   "Carrier_51_G120DStatusWord.0" AT %I2912.0 : Bool;   // Bit_00_READY_RUN
   "Carrier_51_G120DStatusWord.1" AT %I2912.1 : Bool;   // Bit_01_READY_ON
   "Carrier_51_G120DStatusWord.2" AT %I2912.2 : Bool;   // Bit_02_ENABLE
   "Carrier_51_G120DStatusWord.3" AT %I2912.3 : Bool;   // Bit_03_FAULT
   "Carrier_51_G120DStatusWord.4" AT %I2912.4 : Bool;   // Bit_04_OFF2
   "Carrier_51_G120DStatusWord.5" AT %I2912.5 : Bool;   // Bit_05_OFF3
   "Carrier_51_G120DStatusWord.6" AT %I2912.6 : Bool;   // Bit_06_LOCK_OUT
   "Carrier_51_G120DStatusWord.7" AT %I2912.7 : Bool;   // Bit_07_WARN
   "Carrier_51_G120DStatusWord.8" AT %I2913.0 : Bool;   // Bit_08_NO_DEVIATION
   "Carrier_51_G120DStatusWord.9" AT %I2913.1 : Bool;   // Bit_09_CONTR_PLC
   "Carrier_51_G120DStatusWord.10" AT %I2913.2 : Bool;   // Bit_10_F_MAX
   "Carrier_51_G120DStatusWord.11" AT %I2913.3 : Bool;   // Bit_11_LIMIT_REACHED
   "Carrier_51_G120DStatusWord.12" AT %I2913.4 : Bool;   // Bit_12_BRAKE_OPEN
   "Carrier_51_G120DStatusWord.13" AT %I2913.5 : Bool;   // Bit_13_NO_OVERTEMP
   "Carrier_51_G120DStatusWord.14" AT %I2913.6 : Bool;   // Bit_14_CW_CCW
   "Carrier_51_G120DStatusWord.15" AT %I2913.7 : Bool;   // Bit_15_OVERL
   "Carrier_51_Slot2_Input" AT %IW2914 : Word;   // SLOT 2 INPUT WORD
   "Carrier_51_CrashDetectSW" AT %I2914.0 : Bool;   // CRASH DETECT SW
   "Carrier_51_SpareSafetyInput(2_1)" AT %I2914.1 : Bool;   // SPARE SAFETY INPUT
   "Carrier_51_SpareSafetyInput(2_2)" AT %I2914.2 : Bool;   // SPARE SAFETY INPUT
   "Carrier_51_SpareSafetyInput(2_3)" AT %I2914.3 : Bool;   // SPARE SAFETY INPUT
   "Carrier_51_SpareSafetyInput(2_4)" AT %I2914.4 : Bool;   // SPARE SAFETY INPUT
   "Carrier_51_SpareSafetyInput(2_5)" AT %I2914.5 : Bool;   // SPARE SAFETY INPUT
   "Carrier_51_SpareSafetyInput(2_6)" AT %I2914.6 : Bool;   // SPARE SAFETY INPUT
   "Carrier_51_SpareSafetyInput(2_7)" AT %I2914.7 : Bool;   // SPARE SAFETY INPUT
   "Carrier_51_Slot3_SafetyOutput" AT %IW2915 : Word;   // SLOT 3 SAFETY OUTPUT WORD
   "Carrier_51_Crash_Detect_OK" AT %I2915.0 : Bool;   // CARRIER CRASH DETECT
   "Carrier_51_SpareSafetyOutput(3_1)" AT %I2915.1 : Bool;   // SPARE SAFETY OUTPUT
   "Carrier_51_SpareSafetyOutput(3_2)" AT %I2915.2 : Bool;   // SPARE SAFETY OUTPUT
   "Carrier_51_SpareSafetyOutput(3_3)" AT %I2915.3 : Bool;   // SPARE SAFETY OUTPUT
   "Carrier_51_SpareSafetyOutput(3_4)" AT %I2915.4 : Bool;   // SPARE SAFETY OUTPUT
   "Carrier_51_SpareSafetyOutput(3_5)" AT %I2915.5 : Bool;   // SPARE SAFETY OUTPUT
   "Carrier_51_SpareSafetyOutput(3_6)" AT %I2915.6 : Bool;   // SPARE SAFETY OUTPUT
   "Carrier_51_SpareSafetyOutput(3_7)" AT %I2915.7 : Bool;   // SPARE SAFETY OUTPUT
   "Carrier_51_Slot4_Input" AT %IW2916 : Word;   // SLOT 4 INPUT WORD
   "Carrier_51_480VPowerOn_MDCB1" AT %I2916.0 : Bool;   // 480 VAC POWER ON MDCB 1
   "Carrier_51_SpareInput(4_1)" AT %I2916.1 : Bool;   // SPARE INPUT
   "Carrier_51_SpareInput(4_2)" AT %I2916.2 : Bool;   // SPARE INPUT
   "Carrier_51_SitopSelectStatus" AT %I2916.3 : Bool;   // SITOP SELECT STATUS
   "Carrier_51_DCsupplyOnPSCB2" AT %I2916.4 : Bool;   // DC SUPPLY ON PSCB 2
   "Carrier_51_SpareInput(4_5)" AT %I2916.5 : Bool;   // SPARE INPUT
   "Carrier_51_SpareInput(4_6)" AT %I2916.6 : Bool;   // SPARE INPUT
   "Carrier_51_SpareInput(4_7)" AT %I2916.7 : Bool;   // SPARE INPUT
   "Carrier_51_PB1_ProdHoldLH" AT %I2917.0 : Bool;   // PB 1 PRODUCTION HOLD LH
   "Carrier_51_PB2_ResetLH" AT %I2917.1 : Bool;   // PB 2 RESET LH
   "Carrier_51_PB3_ProdHoldRH" AT %I2917.2 : Bool;   // PB 3 PRODUCTION HOLD RH
   "Carrier_51_PB4_ResetRH" AT %I2917.3 : Bool;   // PB 4 RESET RH
   "Carrier_51_SpareInput(4_14)" AT %I2917.4 : Bool;   // SPARE INPUT
   "Carrier_51_SpareInput(4_15)" AT %I2917.5 : Bool;   // SPARE INPUT
   "Carrier_51_SpareInput(4_16)" AT %I2917.6 : Bool;   // SPARE INPUT
   "Carrier_51_SpareInput(4_17)" AT %I2917.7 : Bool;   // SPARE INPUT
   "Carrier_51_Slot5_Output" AT %IW2918 : Word;   // SLOT 5 OUTPUT WORD
   "Carrier_51_IRD400_HMI_24VDC_ENABLE" AT %I2918.0 : Bool;   // IRD 400 PANEL HMI 24V DC POWER
   "Carrier_51_FaultLight_LH" AT %I2918.1 : Bool;   // FAULT LIGHT LH
   "Carrier_51_RunLight_LH" AT %I2918.2 : Bool;   // RUN LIGHT LH
   "Carrier_51_FaultLight_RH" AT %I2918.3 : Bool;   // FAULT LIGHT RH
   "Carrier_51_RunLight_RH" AT %I2918.4 : Bool;   // RUN LIGHT RH
   "Carrier_51_SpareOutput(5_5)" AT %I2918.5 : Bool;   // SPARE OUTPUT
   "Carrier_51_SpareOutput(5_6)" AT %I2918.6 : Bool;   // SPARE OUTPUT
   "Carrier_51_SpareOutput(5_7)" AT %I2918.7 : Bool;   // SPARE OUTPUT
   "Carrier_51_ActualSpeed" AT %IW2920 : Word;   // ACTUAL SPEED
   "Carrier_51_CarrierDriveAlarm" AT %IW2922 : Word;   // CARRIER DRIVE ALARM
   "Carrier_51_CarrierDriveWarning" AT %IW2924 : Word;   // CARRIER DRIVE WARNING
   "Carrier_52_Status" AT %IW2950 : Word;   // CARRIER STATUS WORD
   "Carrier_52_Status.0" AT %I2950.0 : Bool;   // HEARTBEAT
   "Carrier_52_Status.1" AT %I2950.1 : Bool;   // MANUAL
   "Carrier_52_Status.2" AT %I2950.2 : Bool;   // IN_AUTO
   "Carrier_52_Status.3" AT %I2950.3 : Bool;   // POSITIONING_COMPLETE
   "Carrier_52_Status.4" AT %I2950.4 : Bool;   // PRODUCTION HOLD
   "Carrier_52_Status.5" AT %I2950.5 : Bool;   // CARRIER MOVING FORWARD
   "Carrier_52_Status.6" AT %I2950.6 : Bool;   // CARRIER MOVING REVERSE
   "Carrier_52_Status.7" AT %I2950.7 : Bool;   // CARRIER FAULT
   "Carrier_52_Status.8" AT %I2951.0 : Bool;   // CRASH DETECT TRIPPED
   "Carrier_52_Status.9" AT %I2951.1 : Bool;
   "Carrier_52_Status.10" AT %I2951.2 : Bool;
   "Carrier_52_Status.11" AT %I2951.3 : Bool;
   "Carrier_52_Status.12" AT %I2951.4 : Bool;
   "Carrier_52_Status.13" AT %I2951.5 : Bool;
   "Carrier_52_Status.14" AT %I2951.6 : Bool;
   "Carrier_52_Status.15" AT %I2951.7 : Bool;
   "Carrier_52_SDCFaultCode" AT %IW2952 : Word;   // SDC FAULT CODE
   "Carrier_52_CarrierPosition" AT %ID2954 : DWord;   // CARRIER POSITION
   "Carrier_52_CarrierNumber" AT %IW2958 : Word;   // CARRIER NUMBER
   "Carrier_52_G120DControlWord" AT %IW2960 : Word;   // G120D_STW1_CONTROL
   "Carrier_52_G120DControlWord.0" AT %I2960.0 : Bool;   // Bit_00_ON
   "Carrier_52_G120DControlWord.1" AT %I2960.1 : Bool;   // Bit_01_AUS2_INH
   "Carrier_52_G120DControlWord.2" AT %I2960.2 : Bool;   // Bit_02_AUS3_STOP
   "Carrier_52_G120DControlWord.3" AT %I2960.3 : Bool;   // Bit_03_EN
   "Carrier_52_G120DControlWord.4" AT %I2960.4 : Bool;   // Bit_04_EN_RAMP
   "Carrier_52_G120DControlWord.5" AT %I2960.5 : Bool;   // Bit_05_START_RAMP
   "Carrier_52_G120DControlWord.6" AT %I2960.6 : Bool;   // Bit_06_SETPOINT
   "Carrier_52_G120DControlWord.7" AT %I2960.7 : Bool;   // Bit_07_RESET
   "Carrier_52_G120DControlWord.8" AT %I2961.0 : Bool;   // Bit_08_JOG_R
   "Carrier_52_G120DControlWord.9" AT %I2961.1 : Bool;   // Bit_09_JOG_L
   "Carrier_52_G120DControlWord.10" AT %I2961.2 : Bool;   // Bit_10_CONTR_PLC
   "Carrier_52_G120DControlWord.11" AT %I2961.3 : Bool;   // Bit_11_REVERSE
   "Carrier_52_G120DControlWord.12" AT %I2961.4 : Bool;   // Bit_12_BRAKE_RELEASE
   "Carrier_52_G120DControlWord.13" AT %I2961.5 : Bool;   // Bit_13_DDS
   "Carrier_52_G120DControlWord.14" AT %I2961.6 : Bool;   // Bit_14_DO0
   "Carrier_52_G120DControlWord.15" AT %I2961.7 : Bool;   // Bit_15_DO1
   "Carrier_52_G120DStatusWord" AT %IW2962 : Word;   // G120D_ZSW1_STATUS
   "Carrier_52_G120DStatusWord.0" AT %I2962.0 : Bool;   // Bit_00_READY_RUN
   "Carrier_52_G120DStatusWord.1" AT %I2962.1 : Bool;   // Bit_01_READY_ON
   "Carrier_52_G120DStatusWord.2" AT %I2962.2 : Bool;   // Bit_02_ENABLE
   "Carrier_52_G120DStatusWord.3" AT %I2962.3 : Bool;   // Bit_03_FAULT
   "Carrier_52_G120DStatusWord.4" AT %I2962.4 : Bool;   // Bit_04_OFF2
   "Carrier_52_G120DStatusWord.5" AT %I2962.5 : Bool;   // Bit_05_OFF3
   "Carrier_52_G120DStatusWord.6" AT %I2962.6 : Bool;   // Bit_06_LOCK_OUT
   "Carrier_52_G120DStatusWord.7" AT %I2962.7 : Bool;   // Bit_07_WARN
   "Carrier_52_G120DStatusWord.8" AT %I2963.0 : Bool;   // Bit_08_NO_DEVIATION
   "Carrier_52_G120DStatusWord.9" AT %I2963.1 : Bool;   // Bit_09_CONTR_PLC
   "Carrier_52_G120DStatusWord.10" AT %I2963.2 : Bool;   // Bit_10_F_MAX
   "Carrier_52_G120DStatusWord.11" AT %I2963.3 : Bool;   // Bit_11_LIMIT_REACHED
   "Carrier_52_G120DStatusWord.12" AT %I2963.4 : Bool;   // Bit_12_BRAKE_OPEN
   "Carrier_52_G120DStatusWord.13" AT %I2963.5 : Bool;   // Bit_13_NO_OVERTEMP
   "Carrier_52_G120DStatusWord.14" AT %I2963.6 : Bool;   // Bit_14_CW_CCW
   "Carrier_52_G120DStatusWord.15" AT %I2963.7 : Bool;   // Bit_15_OVERL
   "Carrier_52_Slot2_Input" AT %IW2964 : Word;   // SLOT 2 INPUT WORD
   "Carrier_52_CrashDetectSW" AT %I2964.0 : Bool;   // CRASH DETECT SW
   "Carrier_52_SpareSafetyInput(2_1)" AT %I2964.1 : Bool;   // SPARE SAFETY INPUT
   "Carrier_52_SpareSafetyInput(2_2)" AT %I2964.2 : Bool;   // SPARE SAFETY INPUT
   "Carrier_52_SpareSafetyInput(2_3)" AT %I2964.3 : Bool;   // SPARE SAFETY INPUT
   "Carrier_52_SpareSafetyInput(2_4)" AT %I2964.4 : Bool;   // SPARE SAFETY INPUT
   "Carrier_52_SpareSafetyInput(2_5)" AT %I2964.5 : Bool;   // SPARE SAFETY INPUT
   "Carrier_52_SpareSafetyInput(2_6)" AT %I2964.6 : Bool;   // SPARE SAFETY INPUT
   "Carrier_52_SpareSafetyInput(2_7)" AT %I2964.7 : Bool;   // SPARE SAFETY INPUT
   "Carrier_52_Slot3_SafetyOutput" AT %IW2965 : Word;   // SLOT 3 SAFETY OUTPUT WORD
   "Carrier_52_Crash_Detect_OK" AT %I2965.0 : Bool;   // CARRIER CRASH DETECT
   "Carrier_52_SpareSafetyOutput(3_1)" AT %I2965.1 : Bool;   // SPARE SAFETY OUTPUT
   "Carrier_52_SpareSafetyOutput(3_2)" AT %I2965.2 : Bool;   // SPARE SAFETY OUTPUT
   "Carrier_52_SpareSafetyOutput(3_3)" AT %I2965.3 : Bool;   // SPARE SAFETY OUTPUT
   "Carrier_52_SpareSafetyOutput(3_4)" AT %I2965.4 : Bool;   // SPARE SAFETY OUTPUT
   "Carrier_52_SpareSafetyOutput(3_5)" AT %I2965.5 : Bool;   // SPARE SAFETY OUTPUT
   "Carrier_52_SpareSafetyOutput(3_6)" AT %I2965.6 : Bool;   // SPARE SAFETY OUTPUT
   "Carrier_52_SpareSafetyOutput(3_7)" AT %I2965.7 : Bool;   // SPARE SAFETY OUTPUT
   "Carrier_52_Slot4_Input" AT %IW2966 : Word;   // SLOT 4 INPUT WORD
   "Carrier_52_480VPowerOn_MDCB1" AT %I2966.0 : Bool;   // 480 VAC POWER ON MDCB 1
   "Carrier_52_SpareInput(4_1)" AT %I2966.1 : Bool;   // SPARE INPUT
   "Carrier_52_SpareInput(4_2)" AT %I2966.2 : Bool;   // SPARE INPUT
   "Carrier_52_SitopSelectStatus" AT %I2966.3 : Bool;   // SITOP SELECT STATUS
   "Carrier_52_DCsupplyOnPSCB2" AT %I2966.4 : Bool;   // DC SUPPLY ON PSCB 2
   "Carrier_52_SpareInput(4_5)" AT %I2966.5 : Bool;   // SPARE INPUT
   "Carrier_52_SpareInput(4_6)" AT %I2966.6 : Bool;   // SPARE INPUT
   "Carrier_52_SpareInput(4_7)" AT %I2966.7 : Bool;   // SPARE INPUT
   "Carrier_52_PB1_ProdHoldLH" AT %I2967.0 : Bool;   // PB 1 PRODUCTION HOLD LH
   "Carrier_52_PB2_ResetLH" AT %I2967.1 : Bool;   // PB 2 RESET LH
   "Carrier_52_PB3_ProdHoldRH" AT %I2967.2 : Bool;   // PB 3 PRODUCTION HOLD RH
   "Carrier_52_PB4_ResetRH" AT %I2967.3 : Bool;   // PB 4 RESET RH
   "Carrier_52_SpareInput(4_14)" AT %I2967.4 : Bool;   // SPARE INPUT
   "Carrier_52_SpareInput(4_15)" AT %I2967.5 : Bool;   // SPARE INPUT
   "Carrier_52_SpareInput(4_16)" AT %I2967.6 : Bool;   // SPARE INPUT
   "Carrier_52_SpareInput(4_17)" AT %I2967.7 : Bool;   // SPARE INPUT
   "Carrier_52_Slot5_Output" AT %IW2968 : Word;   // SLOT 5 OUTPUT WORD
   "Carrier_52_IRD400_HMI_24VDC_ENABLE" AT %I2968.0 : Bool;   // IRD 400 PANEL HMI 24V DC POWER
   "Carrier_52_FaultLight_LH" AT %I2968.1 : Bool;   // FAULT LIGHT LH
   "Carrier_52_RunLight_LH" AT %I2968.2 : Bool;   // RUN LIGHT LH
   "Carrier_52_FaultLight_RH" AT %I2968.3 : Bool;   // FAULT LIGHT RH
   "Carrier_52_RunLight_RH" AT %I2968.4 : Bool;   // RUN LIGHT RH
   "Carrier_52_SpareOutput(5_5)" AT %I2968.5 : Bool;   // SPARE OUTPUT
   "Carrier_52_SpareOutput(5_6)" AT %I2968.6 : Bool;   // SPARE OUTPUT
   "Carrier_52_SpareOutput(5_7)" AT %I2968.7 : Bool;   // SPARE OUTPUT
   "Carrier_52_ActualSpeed" AT %IW2970 : Word;   // ACTUAL SPEED
   "Carrier_52_CarrierDriveAlarm" AT %IW2972 : Word;   // CARRIER DRIVE ALARM
   "Carrier_52_CarrierDriveWarning" AT %IW2974 : Word;   // CARRIER DRIVE WARNING
   "Carrier_53_Status" AT %IW3000 : Word;   // CARRIER STATUS WORD
   "Carrier_53_Status.0" AT %I3000.0 : Bool;   // HEARTBEAT
   "Carrier_53_Status.1" AT %I3000.1 : Bool;   // MANUAL
   "Carrier_53_Status.2" AT %I3000.2 : Bool;   // IN_AUTO
   "Carrier_53_Status.3" AT %I3000.3 : Bool;   // POSITIONING_COMPLETE
   "Carrier_53_Status.4" AT %I3000.4 : Bool;   // PRODUCTION HOLD
   "Carrier_53_Status.5" AT %I3000.5 : Bool;   // CARRIER MOVING FORWARD
   "Carrier_53_Status.6" AT %I3000.6 : Bool;   // CARRIER MOVING REVERSE
   "Carrier_53_Status.7" AT %I3000.7 : Bool;   // CARRIER FAULT
   "Carrier_53_Status.8" AT %I3001.0 : Bool;   // CRASH DETECT TRIPPED
   "Carrier_53_Status.9" AT %I3001.1 : Bool;
   "Carrier_53_Status.10" AT %I3001.2 : Bool;
   "Carrier_53_Status.11" AT %I3001.3 : Bool;
   "Carrier_53_Status.12" AT %I3001.4 : Bool;
   "Carrier_53_Status.13" AT %I3001.5 : Bool;
   "Carrier_53_Status.14" AT %I3001.6 : Bool;
   "Carrier_53_Status.15" AT %I3001.7 : Bool;
   "Carrier_53_SDCFaultCode" AT %IW3002 : Word;   // SDC FAULT CODE
   "Carrier_53_CarrierPosition" AT %ID3004 : DWord;   // CARRIER POSITION
   "Carrier_53_CarrierNumber" AT %IW3008 : Word;   // CARRIER NUMBER
   "Carrier_53_G120DControlWord" AT %IW3010 : Word;   // G120D_STW1_CONTROL
   "Carrier_53_G120DControlWord.0" AT %I3010.0 : Bool;   // Bit_00_ON
   "Carrier_53_G120DControlWord.1" AT %I3010.1 : Bool;   // Bit_01_AUS2_INH
   "Carrier_53_G120DControlWord.2" AT %I3010.2 : Bool;   // Bit_02_AUS3_STOP
   "Carrier_53_G120DControlWord.3" AT %I3010.3 : Bool;   // Bit_03_EN
   "Carrier_53_G120DControlWord.4" AT %I3010.4 : Bool;   // Bit_04_EN_RAMP
   "Carrier_53_G120DControlWord.5" AT %I3010.5 : Bool;   // Bit_05_START_RAMP
   "Carrier_53_G120DControlWord.6" AT %I3010.6 : Bool;   // Bit_06_SETPOINT
   "Carrier_53_G120DControlWord.7" AT %I3010.7 : Bool;   // Bit_07_RESET
   "Carrier_53_G120DControlWord.8" AT %I3011.0 : Bool;   // Bit_08_JOG_R
   "Carrier_53_G120DControlWord.9" AT %I3011.1 : Bool;   // Bit_09_JOG_L
   "Carrier_53_G120DControlWord.10" AT %I3011.2 : Bool;   // Bit_10_CONTR_PLC
   "Carrier_53_G120DControlWord.11" AT %I3011.3 : Bool;   // Bit_11_REVERSE
   "Carrier_53_G120DControlWord.12" AT %I3011.4 : Bool;   // Bit_12_BRAKE_RELEASE
   "Carrier_53_G120DControlWord.13" AT %I3011.5 : Bool;   // Bit_13_DDS
   "Carrier_53_G120DControlWord.14" AT %I3011.6 : Bool;   // Bit_14_DO0
   "Carrier_53_G120DControlWord.15" AT %I3011.7 : Bool;   // Bit_15_DO1
   "Carrier_53_G120DStatusWord" AT %IW3012 : Word;   // G120D_ZSW1_STATUS
   "Carrier_53_G120DStatusWord.0" AT %I3012.0 : Bool;   // Bit_00_READY_RUN
   "Carrier_53_G120DStatusWord.1" AT %I3012.1 : Bool;   // Bit_01_READY_ON
   "Carrier_53_G120DStatusWord.2" AT %I3012.2 : Bool;   // Bit_02_ENABLE
   "Carrier_53_G120DStatusWord.3" AT %I3012.3 : Bool;   // Bit_03_FAULT
   "Carrier_53_G120DStatusWord.4" AT %I3012.4 : Bool;   // Bit_04_OFF2
   "Carrier_53_G120DStatusWord.5" AT %I3012.5 : Bool;   // Bit_05_OFF3
   "Carrier_53_G120DStatusWord.6" AT %I3012.6 : Bool;   // Bit_06_LOCK_OUT
   "Carrier_53_G120DStatusWord.7" AT %I3012.7 : Bool;   // Bit_07_WARN
   "Carrier_53_G120DStatusWord.8" AT %I3013.0 : Bool;   // Bit_08_NO_DEVIATION
   "Carrier_53_G120DStatusWord.9" AT %I3013.1 : Bool;   // Bit_09_CONTR_PLC
   "Carrier_53_G120DStatusWord.10" AT %I3013.2 : Bool;   // Bit_10_F_MAX
   "Carrier_53_G120DStatusWord.11" AT %I3013.3 : Bool;   // Bit_11_LIMIT_REACHED
   "Carrier_53_G120DStatusWord.12" AT %I3013.4 : Bool;   // Bit_12_BRAKE_OPEN
   "Carrier_53_G120DStatusWord.13" AT %I3013.5 : Bool;   // Bit_13_NO_OVERTEMP
   "Carrier_53_G120DStatusWord.14" AT %I3013.6 : Bool;   // Bit_14_CW_CCW
   "Carrier_53_G120DStatusWord.15" AT %I3013.7 : Bool;   // Bit_15_OVERL
   "Carrier_53_Slot2_Input" AT %IW3014 : Word;   // SLOT 2 INPUT WORD
   "Carrier_53_CrashDetectSW" AT %I3014.0 : Bool;   // CRASH DETECT SW
   "Carrier_53_SpareSafetyInput(2_1)" AT %I3014.1 : Bool;   // SPARE SAFETY INPUT
   "Carrier_53_SpareSafetyInput(2_2)" AT %I3014.2 : Bool;   // SPARE SAFETY INPUT
   "Carrier_53_SpareSafetyInput(2_3)" AT %I3014.3 : Bool;   // SPARE SAFETY INPUT
   "Carrier_53_SpareSafetyInput(2_4)" AT %I3014.4 : Bool;   // SPARE SAFETY INPUT
   "Carrier_53_SpareSafetyInput(2_5)" AT %I3014.5 : Bool;   // SPARE SAFETY INPUT
   "Carrier_53_SpareSafetyInput(2_6)" AT %I3014.6 : Bool;   // SPARE SAFETY INPUT
   "Carrier_53_SpareSafetyInput(2_7)" AT %I3014.7 : Bool;   // SPARE SAFETY INPUT
   "Carrier_53_Slot3_SafetyOutput" AT %IW3015 : Word;   // SLOT 3 SAFETY OUTPUT WORD
   "Carrier_53_Crash_Detect_OK" AT %I3015.0 : Bool;   // CARRIER CRASH DETECT
   "Carrier_53_SpareSafetyOutput(3_1)" AT %I3015.1 : Bool;   // SPARE SAFETY OUTPUT
   "Carrier_53_SpareSafetyOutput(3_2)" AT %I3015.2 : Bool;   // SPARE SAFETY OUTPUT
   "Carrier_53_SpareSafetyOutput(3_3)" AT %I3015.3 : Bool;   // SPARE SAFETY OUTPUT
   "Carrier_53_SpareSafetyOutput(3_4)" AT %I3015.4 : Bool;   // SPARE SAFETY OUTPUT
   "Carrier_53_SpareSafetyOutput(3_5)" AT %I3015.5 : Bool;   // SPARE SAFETY OUTPUT
   "Carrier_53_SpareSafetyOutput(3_6)" AT %I3015.6 : Bool;   // SPARE SAFETY OUTPUT
   "Carrier_53_SpareSafetyOutput(3_7)" AT %I3015.7 : Bool;   // SPARE SAFETY OUTPUT
   "Carrier_53_Slot4_Input" AT %IW3016 : Word;   // SLOT 4 INPUT WORD
   "Carrier_53_480VPowerOn_MDCB1" AT %I3016.0 : Bool;   // 480 VAC POWER ON MDCB 1
   "Carrier_53_SpareInput(4_1)" AT %I3016.1 : Bool;   // SPARE INPUT
   "Carrier_53_SpareInput(4_2)" AT %I3016.2 : Bool;   // SPARE INPUT
   "Carrier_53_SitopSelectStatus" AT %I3016.3 : Bool;   // SITOP SELECT STATUS
   "Carrier_53_DCsupplyOnPSCB2" AT %I3016.4 : Bool;   // DC SUPPLY ON PSCB 2
   "Carrier_53_SpareInput(4_5)" AT %I3016.5 : Bool;   // SPARE INPUT
   "Carrier_53_SpareInput(4_6)" AT %I3016.6 : Bool;   // SPARE INPUT
   "Carrier_53_SpareInput(4_7)" AT %I3016.7 : Bool;   // SPARE INPUT
   "Carrier_53_PB1_ProdHoldLH" AT %I3017.0 : Bool;   // PB 1 PRODUCTION HOLD LH
   "Carrier_53_PB2_ResetLH" AT %I3017.1 : Bool;   // PB 2 RESET LH
   "Carrier_53_PB3_ProdHoldRH" AT %I3017.2 : Bool;   // PB 3 PRODUCTION HOLD RH
   "Carrier_53_PB4_ResetRH" AT %I3017.3 : Bool;   // PB 4 RESET RH
   "Carrier_53_SpareInput(4_14)" AT %I3017.4 : Bool;   // SPARE INPUT
   "Carrier_53_SpareInput(4_15)" AT %I3017.5 : Bool;   // SPARE INPUT
   "Carrier_53_SpareInput(4_16)" AT %I3017.6 : Bool;   // SPARE INPUT
   "Carrier_53_SpareInput(4_17)" AT %I3017.7 : Bool;   // SPARE INPUT
   "Carrier_53_Slot5_Output" AT %IW3018 : Word;   // SLOT 5 OUTPUT WORD
   "Carrier_53_IRD400_HMI_24VDC_ENABLE" AT %I3018.0 : Bool;   // IRD 400 PANEL HMI 24V DC POWER
   "Carrier_53_FaultLight_LH" AT %I3018.1 : Bool;   // FAULT LIGHT LH
   "Carrier_53_RunLight_LH" AT %I3018.2 : Bool;   // RUN LIGHT LH
   "Carrier_53_FaultLight_RH" AT %I3018.3 : Bool;   // FAULT LIGHT RH
   "Carrier_53_RunLight_RH" AT %I3018.4 : Bool;   // RUN LIGHT RH
   "Carrier_53_SpareOutput(5_5)" AT %I3018.5 : Bool;   // SPARE OUTPUT
   "Carrier_53_SpareOutput(5_6)" AT %I3018.6 : Bool;   // SPARE OUTPUT
   "Carrier_53_SpareOutput(5_7)" AT %I3018.7 : Bool;   // SPARE OUTPUT
   "Carrier_53_ActualSpeed" AT %IW3020 : Word;   // ACTUAL SPEED
   "Carrier_53_CarrierDriveAlarm" AT %IW3022 : Word;   // CARRIER DRIVE ALARM
   "Carrier_53_CarrierDriveWarning" AT %IW3024 : Word;   // CARRIER DRIVE WARNING
   "Carrier_54_Status" AT %IW3050 : Word;   // CARRIER STATUS WORD
   "Carrier_54_Status.0" AT %I3050.0 : Bool;   // HEARTBEAT
   "Carrier_54_Status.1" AT %I3050.1 : Bool;   // MANUAL
   "Carrier_54_Status.2" AT %I3050.2 : Bool;   // IN_AUTO
   "Carrier_54_Status.3" AT %I3050.3 : Bool;   // POSITIONING_COMPLETE
   "Carrier_54_Status.4" AT %I3050.4 : Bool;   // PRODUCTION HOLD
   "Carrier_54_Status.5" AT %I3050.5 : Bool;   // CARRIER MOVING FORWARD
   "Carrier_54_Status.6" AT %I3050.6 : Bool;   // CARRIER MOVING REVERSE
   "Carrier_54_Status.7" AT %I3050.7 : Bool;   // CARRIER FAULT
   "Carrier_54_Status.8" AT %I3051.0 : Bool;   // CRASH DETECT TRIPPED
   "Carrier_54_Status.9" AT %I3051.1 : Bool;
   "Carrier_54_Status.10" AT %I3051.2 : Bool;
   "Carrier_54_Status.11" AT %I3051.3 : Bool;
   "Carrier_54_Status.12" AT %I3051.4 : Bool;
   "Carrier_54_Status.13" AT %I3051.5 : Bool;
   "Carrier_54_Status.14" AT %I3051.6 : Bool;
   "Carrier_54_Status.15" AT %I3051.7 : Bool;
   "Carrier_54_SDCFaultCode" AT %IW3052 : Word;   // SDC FAULT CODE
   "Carrier_54_CarrierPosition" AT %ID3054 : DWord;   // CARRIER POSITION
   "Carrier_54_CarrierNumber" AT %IW3058 : Word;   // CARRIER NUMBER
   "Carrier_54_G120DControlWord" AT %IW3060 : Word;   // G120D_STW1_CONTROL
   "Carrier_54_G120DControlWord.0" AT %I3060.0 : Bool;   // Bit_00_ON
   "Carrier_54_G120DControlWord.1" AT %I3060.1 : Bool;   // Bit_01_AUS2_INH
   "Carrier_54_G120DControlWord.2" AT %I3060.2 : Bool;   // Bit_02_AUS3_STOP
   "Carrier_54_G120DControlWord.3" AT %I3060.3 : Bool;   // Bit_03_EN
   "Carrier_54_G120DControlWord.4" AT %I3060.4 : Bool;   // Bit_04_EN_RAMP
   "Carrier_54_G120DControlWord.5" AT %I3060.5 : Bool;   // Bit_05_START_RAMP
   "Carrier_54_G120DControlWord.6" AT %I3060.6 : Bool;   // Bit_06_SETPOINT
   "Carrier_54_G120DControlWord.7" AT %I3060.7 : Bool;   // Bit_07_RESET
   "Carrier_54_G120DControlWord.8" AT %I3061.0 : Bool;   // Bit_08_JOG_R
   "Carrier_54_G120DControlWord.9" AT %I3061.1 : Bool;   // Bit_09_JOG_L
   "Carrier_54_G120DControlWord.10" AT %I3061.2 : Bool;   // Bit_10_CONTR_PLC
   "Carrier_54_G120DControlWord.11" AT %I3061.3 : Bool;   // Bit_11_REVERSE
   "Carrier_54_G120DControlWord.12" AT %I3061.4 : Bool;   // Bit_12_BRAKE_RELEASE
   "Carrier_54_G120DControlWord.13" AT %I3061.5 : Bool;   // Bit_13_DDS
   "Carrier_54_G120DControlWord.14" AT %I3061.6 : Bool;   // Bit_14_DO0
   "Carrier_54_G120DControlWord.15" AT %I3061.7 : Bool;   // Bit_15_DO1
   "Carrier_54_G120DStatusWord" AT %IW3062 : Word;   // G120D_ZSW1_STATUS
   "Carrier_54_G120DStatusWord.0" AT %I3062.0 : Bool;   // Bit_00_READY_RUN
   "Carrier_54_G120DStatusWord.1" AT %I3062.1 : Bool;   // Bit_01_READY_ON
   "Carrier_54_G120DStatusWord.2" AT %I3062.2 : Bool;   // Bit_02_ENABLE
   "Carrier_54_G120DStatusWord.3" AT %I3062.3 : Bool;   // Bit_03_FAULT
   "Carrier_54_G120DStatusWord.4" AT %I3062.4 : Bool;   // Bit_04_OFF2
   "Carrier_54_G120DStatusWord.5" AT %I3062.5 : Bool;   // Bit_05_OFF3
   "Carrier_54_G120DStatusWord.6" AT %I3062.6 : Bool;   // Bit_06_LOCK_OUT
   "Carrier_54_G120DStatusWord.7" AT %I3062.7 : Bool;   // Bit_07_WARN
   "Carrier_54_G120DStatusWord.8" AT %I3063.0 : Bool;   // Bit_08_NO_DEVIATION
   "Carrier_54_G120DStatusWord.9" AT %I3063.1 : Bool;   // Bit_09_CONTR_PLC
   "Carrier_54_G120DStatusWord.10" AT %I3063.2 : Bool;   // Bit_10_F_MAX
   "Carrier_54_G120DStatusWord.11" AT %I3063.3 : Bool;   // Bit_11_LIMIT_REACHED
   "Carrier_54_G120DStatusWord.12" AT %I3063.4 : Bool;   // Bit_12_BRAKE_OPEN
   "Carrier_54_G120DStatusWord.13" AT %I3063.5 : Bool;   // Bit_13_NO_OVERTEMP
   "Carrier_54_G120DStatusWord.14" AT %I3063.6 : Bool;   // Bit_14_CW_CCW
   "Carrier_54_G120DStatusWord.15" AT %I3063.7 : Bool;   // Bit_15_OVERL
   "Carrier_54_Slot2_Input" AT %IW3064 : Word;   // SLOT 2 INPUT WORD
   "Carrier_54_CrashDetectSW" AT %I3064.0 : Bool;   // CRASH DETECT SW
   "Carrier_54_SpareSafetyInput(2_1)" AT %I3064.1 : Bool;   // SPARE SAFETY INPUT
   "Carrier_54_SpareSafetyInput(2_2)" AT %I3064.2 : Bool;   // SPARE SAFETY INPUT
   "Carrier_54_SpareSafetyInput(2_3)" AT %I3064.3 : Bool;   // SPARE SAFETY INPUT
   "Carrier_54_SpareSafetyInput(2_4)" AT %I3064.4 : Bool;   // SPARE SAFETY INPUT
   "Carrier_54_SpareSafetyInput(2_5)" AT %I3064.5 : Bool;   // SPARE SAFETY INPUT
   "Carrier_54_SpareSafetyInput(2_6)" AT %I3064.6 : Bool;   // SPARE SAFETY INPUT
   "Carrier_54_SpareSafetyInput(2_7)" AT %I3064.7 : Bool;   // SPARE SAFETY INPUT
   "Carrier_54_Slot3_SafetyOutput" AT %IW3065 : Word;   // SLOT 3 SAFETY OUTPUT WORD
   "Carrier_54_Crash_Detect_OK" AT %I3065.0 : Bool;   // CARRIER CRASH DETECT
   "Carrier_54_SpareSafetyOutput(3_1)" AT %I3065.1 : Bool;   // SPARE SAFETY OUTPUT
   "Carrier_54_SpareSafetyOutput(3_2)" AT %I3065.2 : Bool;   // SPARE SAFETY OUTPUT
   "Carrier_54_SpareSafetyOutput(3_3)" AT %I3065.3 : Bool;   // SPARE SAFETY OUTPUT
   "Carrier_54_SpareSafetyOutput(3_4)" AT %I3065.4 : Bool;   // SPARE SAFETY OUTPUT
   "Carrier_54_SpareSafetyOutput(3_5)" AT %I3065.5 : Bool;   // SPARE SAFETY OUTPUT
   "Carrier_54_SpareSafetyOutput(3_6)" AT %I3065.6 : Bool;   // SPARE SAFETY OUTPUT
   "Carrier_54_SpareSafetyOutput(3_7)" AT %I3065.7 : Bool;   // SPARE SAFETY OUTPUT
   "Carrier_54_Slot4_Input" AT %IW3066 : Word;   // SLOT 4 INPUT WORD
   "Carrier_54_480VPowerOn_MDCB1" AT %I3066.0 : Bool;   // 480 VAC POWER ON MDCB 1
   "Carrier_54_SpareInput(4_1)" AT %I3066.1 : Bool;   // SPARE INPUT
   "Carrier_54_SpareInput(4_2)" AT %I3066.2 : Bool;   // SPARE INPUT
   "Carrier_54_SitopSelectStatus" AT %I3066.3 : Bool;   // SITOP SELECT STATUS
   "Carrier_54_DCsupplyOnPSCB2" AT %I3066.4 : Bool;   // DC SUPPLY ON PSCB 2
   "Carrier_54_SpareInput(4_5)" AT %I3066.5 : Bool;   // SPARE INPUT
   "Carrier_54_SpareInput(4_6)" AT %I3066.6 : Bool;   // SPARE INPUT
   "Carrier_54_SpareInput(4_7)" AT %I3066.7 : Bool;   // SPARE INPUT
   "Carrier_54_PB1_ProdHoldLH" AT %I3067.0 : Bool;   // PB 1 PRODUCTION HOLD LH
   "Carrier_54_PB2_ResetLH" AT %I3067.1 : Bool;   // PB 2 RESET LH
   "Carrier_54_PB3_ProdHoldRH" AT %I3067.2 : Bool;   // PB 3 PRODUCTION HOLD RH
   "Carrier_54_PB4_ResetRH" AT %I3067.3 : Bool;   // PB 4 RESET RH
   "Carrier_54_SpareInput(4_14)" AT %I3067.4 : Bool;   // SPARE INPUT
   "Carrier_54_SpareInput(4_15)" AT %I3067.5 : Bool;   // SPARE INPUT
   "Carrier_54_SpareInput(4_16)" AT %I3067.6 : Bool;   // SPARE INPUT
   "Carrier_54_SpareInput(4_17)" AT %I3067.7 : Bool;   // SPARE INPUT
   "Carrier_54_Slot5_Output" AT %IW3068 : Word;   // SLOT 5 OUTPUT WORD
   "Carrier_54_IRD400_HMI_24VDC_ENABLE" AT %I3068.0 : Bool;   // IRD 400 PANEL HMI 24V DC POWER
   "Carrier_54_FaultLight_LH" AT %I3068.1 : Bool;   // FAULT LIGHT LH
   "Carrier_54_RunLight_LH" AT %I3068.2 : Bool;   // RUN LIGHT LH
   "Carrier_54_FaultLight_RH" AT %I3068.3 : Bool;   // FAULT LIGHT RH
   "Carrier_54_RunLight_RH" AT %I3068.4 : Bool;   // RUN LIGHT RH
   "Carrier_54_SpareOutput(5_5)" AT %I3068.5 : Bool;   // SPARE OUTPUT
   "Carrier_54_SpareOutput(5_6)" AT %I3068.6 : Bool;   // SPARE OUTPUT
   "Carrier_54_SpareOutput(5_7)" AT %I3068.7 : Bool;   // SPARE OUTPUT
   "Carrier_54_ActualSpeed" AT %IW3070 : Word;   // ACTUAL SPEED
   "Carrier_54_CarrierDriveAlarm" AT %IW3072 : Word;   // CARRIER DRIVE ALARM
   "Carrier_54_CarrierDriveWarning" AT %IW3074 : Word;   // CARRIER DRIVE WARNING
   "Carrier_55_Status" AT %IW3100 : Word;   // CARRIER STATUS WORD
   "Carrier_55_Status.0" AT %I3100.0 : Bool;   // HEARTBEAT
   "Carrier_55_Status.1" AT %I3100.1 : Bool;   // MANUAL
   "Carrier_55_Status.2" AT %I3100.2 : Bool;   // IN_AUTO
   "Carrier_55_Status.3" AT %I3100.3 : Bool;   // POSITIONING_COMPLETE
   "Carrier_55_Status.4" AT %I3100.4 : Bool;   // PRODUCTION HOLD
   "Carrier_55_Status.5" AT %I3100.5 : Bool;   // CARRIER MOVING FORWARD
   "Carrier_55_Status.6" AT %I3100.6 : Bool;   // CARRIER MOVING REVERSE
   "Carrier_55_Status.7" AT %I3100.7 : Bool;   // CARRIER FAULT
   "Carrier_55_Status.8" AT %I3101.0 : Bool;   // CRASH DETECT TRIPPED
   "Carrier_55_Status.9" AT %I3101.1 : Bool;
   "Carrier_55_Status.10" AT %I3101.2 : Bool;
   "Carrier_55_Status.11" AT %I3101.3 : Bool;
   "Carrier_55_Status.12" AT %I3101.4 : Bool;
   "Carrier_55_Status.13" AT %I3101.5 : Bool;
   "Carrier_55_Status.14" AT %I3101.6 : Bool;
   "Carrier_55_Status.15" AT %I3101.7 : Bool;
   "Carrier_55_SDCFaultCode" AT %IW3102 : Word;   // SDC FAULT CODE
   "Carrier_55_CarrierPosition" AT %ID3104 : DWord;   // CARRIER POSITION
   "Carrier_55_CarrierNumber" AT %IW3108 : Word;   // CARRIER NUMBER
   "Carrier_55_G120DControlWord" AT %IW3110 : Word;   // G120D_STW1_CONTROL
   "Carrier_55_G120DControlWord.0" AT %I3110.0 : Bool;   // Bit_00_ON
   "Carrier_55_G120DControlWord.1" AT %I3110.1 : Bool;   // Bit_01_AUS2_INH
   "Carrier_55_G120DControlWord.2" AT %I3110.2 : Bool;   // Bit_02_AUS3_STOP
   "Carrier_55_G120DControlWord.3" AT %I3110.3 : Bool;   // Bit_03_EN
   "Carrier_55_G120DControlWord.4" AT %I3110.4 : Bool;   // Bit_04_EN_RAMP
   "Carrier_55_G120DControlWord.5" AT %I3110.5 : Bool;   // Bit_05_START_RAMP
   "Carrier_55_G120DControlWord.6" AT %I3110.6 : Bool;   // Bit_06_SETPOINT
   "Carrier_55_G120DControlWord.7" AT %I3110.7 : Bool;   // Bit_07_RESET
   "Carrier_55_G120DControlWord.8" AT %I3111.0 : Bool;   // Bit_08_JOG_R
   "Carrier_55_G120DControlWord.9" AT %I3111.1 : Bool;   // Bit_09_JOG_L
   "Carrier_55_G120DControlWord.10" AT %I3111.2 : Bool;   // Bit_10_CONTR_PLC
   "Carrier_55_G120DControlWord.11" AT %I3111.3 : Bool;   // Bit_11_REVERSE
   "Carrier_55_G120DControlWord.12" AT %I3111.4 : Bool;   // Bit_12_BRAKE_RELEASE
   "Carrier_55_G120DControlWord.13" AT %I3111.5 : Bool;   // Bit_13_DDS
   "Carrier_55_G120DControlWord.14" AT %I3111.6 : Bool;   // Bit_14_DO0
   "Carrier_55_G120DControlWord.15" AT %I3111.7 : Bool;   // Bit_15_DO1
   "Carrier_55_G120DStatusWord" AT %IW3112 : Word;   // G120D_ZSW1_STATUS
   "Carrier_55_G120DStatusWord.0" AT %I3112.0 : Bool;   // Bit_00_READY_RUN
   "Carrier_55_G120DStatusWord.1" AT %I3112.1 : Bool;   // Bit_01_READY_ON
   "Carrier_55_G120DStatusWord.2" AT %I3112.2 : Bool;   // Bit_02_ENABLE
   "Carrier_55_G120DStatusWord.3" AT %I3112.3 : Bool;   // Bit_03_FAULT
   "Carrier_55_G120DStatusWord.4" AT %I3112.4 : Bool;   // Bit_04_OFF2
   "Carrier_55_G120DStatusWord.5" AT %I3112.5 : Bool;   // Bit_05_OFF3
   "Carrier_55_G120DStatusWord.6" AT %I3112.6 : Bool;   // Bit_06_LOCK_OUT
   "Carrier_55_G120DStatusWord.7" AT %I3112.7 : Bool;   // Bit_07_WARN
   "Carrier_55_G120DStatusWord.8" AT %I3113.0 : Bool;   // Bit_08_NO_DEVIATION
   "Carrier_55_G120DStatusWord.9" AT %I3113.1 : Bool;   // Bit_09_CONTR_PLC
   "Carrier_55_G120DStatusWord.10" AT %I3113.2 : Bool;   // Bit_10_F_MAX
   "Carrier_55_G120DStatusWord.11" AT %I3113.3 : Bool;   // Bit_11_LIMIT_REACHED
   "Carrier_55_G120DStatusWord.12" AT %I3113.4 : Bool;   // Bit_12_BRAKE_OPEN
   "Carrier_55_G120DStatusWord.13" AT %I3113.5 : Bool;   // Bit_13_NO_OVERTEMP
   "Carrier_55_G120DStatusWord.14" AT %I3113.6 : Bool;   // Bit_14_CW_CCW
   "Carrier_55_G120DStatusWord.15" AT %I3113.7 : Bool;   // Bit_15_OVERL
   "Carrier_55_Slot2_Input" AT %IW3114 : Word;   // SLOT 2 INPUT WORD
   "Carrier_55_CrashDetectSW" AT %I3114.0 : Bool;   // CRASH DETECT SW
   "Carrier_55_SpareSafetyInput(2_1)" AT %I3114.1 : Bool;   // SPARE SAFETY INPUT
   "Carrier_55_SpareSafetyInput(2_2)" AT %I3114.2 : Bool;   // SPARE SAFETY INPUT
   "Carrier_55_SpareSafetyInput(2_3)" AT %I3114.3 : Bool;   // SPARE SAFETY INPUT
   "Carrier_55_SpareSafetyInput(2_4)" AT %I3114.4 : Bool;   // SPARE SAFETY INPUT
   "Carrier_55_SpareSafetyInput(2_5)" AT %I3114.5 : Bool;   // SPARE SAFETY INPUT
   "Carrier_55_SpareSafetyInput(2_6)" AT %I3114.6 : Bool;   // SPARE SAFETY INPUT
   "Carrier_55_SpareSafetyInput(2_7)" AT %I3114.7 : Bool;   // SPARE SAFETY INPUT
   "Carrier_55_Slot3_SafetyOutput" AT %IW3115 : Word;   // SLOT 3 SAFETY OUTPUT WORD
   "Carrier_55_Crash_Detect_OK" AT %I3115.0 : Bool;   // CARRIER CRASH DETECT
   "Carrier_55_SpareSafetyOutput(3_1)" AT %I3115.1 : Bool;   // SPARE SAFETY OUTPUT
   "Carrier_55_SpareSafetyOutput(3_2)" AT %I3115.2 : Bool;   // SPARE SAFETY OUTPUT
   "Carrier_55_SpareSafetyOutput(3_3)" AT %I3115.3 : Bool;   // SPARE SAFETY OUTPUT
   "Carrier_55_SpareSafetyOutput(3_4)" AT %I3115.4 : Bool;   // SPARE SAFETY OUTPUT
   "Carrier_55_SpareSafetyOutput(3_5)" AT %I3115.5 : Bool;   // SPARE SAFETY OUTPUT
   "Carrier_55_SpareSafetyOutput(3_6)" AT %I3115.6 : Bool;   // SPARE SAFETY OUTPUT
   "Carrier_55_SpareSafetyOutput(3_7)" AT %I3115.7 : Bool;   // SPARE SAFETY OUTPUT
   "Carrier_55_Slot4_Input" AT %IW3116 : Word;   // SLOT 4 INPUT WORD
   "Carrier_55_480VPowerOn_MDCB1" AT %I3116.0 : Bool;   // 480 VAC POWER ON MDCB 1
   "Carrier_55_SpareInput(4_1)" AT %I3116.1 : Bool;   // SPARE INPUT
   "Carrier_55_SpareInput(4_2)" AT %I3116.2 : Bool;   // SPARE INPUT
   "Carrier_55_SitopSelectStatus" AT %I3116.3 : Bool;   // SITOP SELECT STATUS
   "Carrier_55_DCsupplyOnPSCB2" AT %I3116.4 : Bool;   // DC SUPPLY ON PSCB 2
   "Carrier_55_SpareInput(4_5)" AT %I3116.5 : Bool;   // SPARE INPUT
   "Carrier_55_SpareInput(4_6)" AT %I3116.6 : Bool;   // SPARE INPUT
   "Carrier_55_SpareInput(4_7)" AT %I3116.7 : Bool;   // SPARE INPUT
   "Carrier_55_PB1_ProdHoldLH" AT %I3117.0 : Bool;   // PB 1 PRODUCTION HOLD LH
   "Carrier_55_PB2_ResetLH" AT %I3117.1 : Bool;   // PB 2 RESET LH
   "Carrier_55_PB3_ProdHoldRH" AT %I3117.2 : Bool;   // PB 3 PRODUCTION HOLD RH
   "Carrier_55_PB4_ResetRH" AT %I3117.3 : Bool;   // PB 4 RESET RH
   "Carrier_55_SpareInput(4_14)" AT %I3117.4 : Bool;   // SPARE INPUT
   "Carrier_55_SpareInput(4_15)" AT %I3117.5 : Bool;   // SPARE INPUT
   "Carrier_55_SpareInput(4_16)" AT %I3117.6 : Bool;   // SPARE INPUT
   "Carrier_55_SpareInput(4_17)" AT %I3117.7 : Bool;   // SPARE INPUT
   "Carrier_55_Slot5_Output" AT %IW3118 : Word;   // SLOT 5 OUTPUT WORD
   "Carrier_55_IRD400_HMI_24VDC_ENABLE" AT %I3118.0 : Bool;   // IRD 400 PANEL HMI 24V DC POWER
